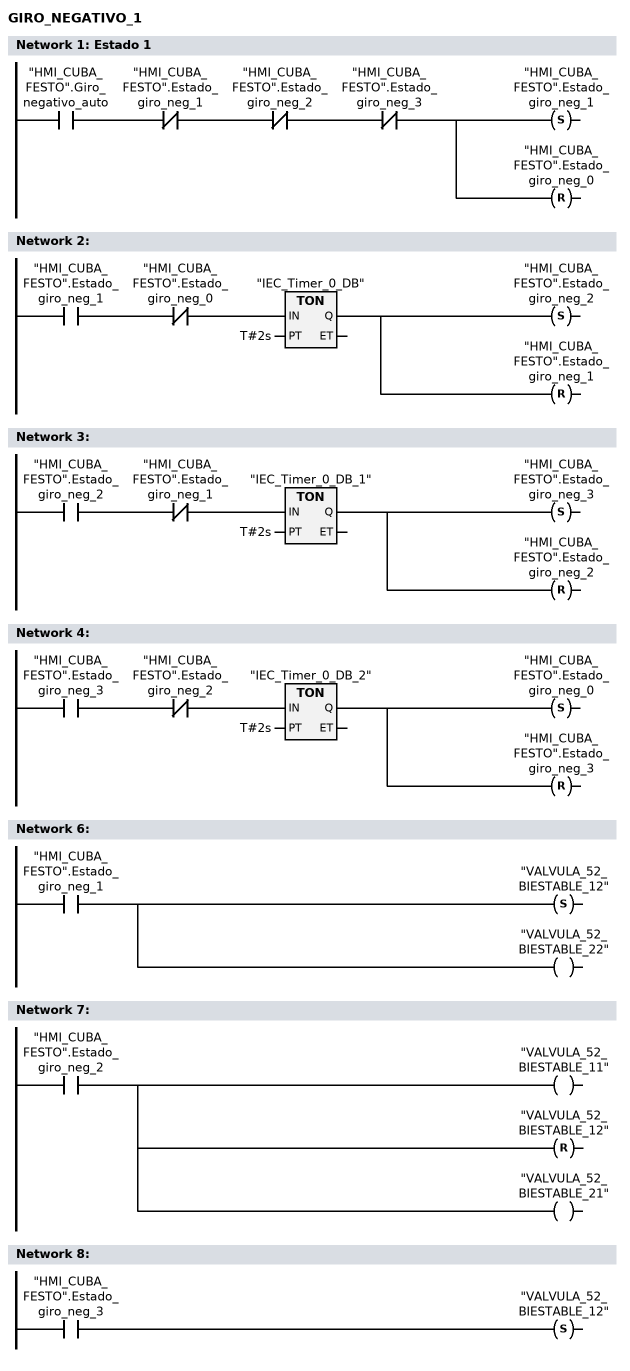
   RUNG wire#powerrail
      Contact( "HMI_CUBA_FESTO".Giro_negativo_auto )
      I_Contact( "HMI_CUBA_FESTO".Estado_giro_neg_1 )
      I_Contact( "HMI_CUBA_FESTO".Estado_giro_neg_2 )
      I_Contact( "HMI_CUBA_FESTO".Estado_giro_neg_3 )
      wire#w1
      S_Coil( "HMI_CUBA_FESTO".Estado_giro_neg_1 )
   END_RUNG
   RUNG wire#w1
      R_Coil( "HMI_CUBA_FESTO".Estado_giro_neg_0 )
   END_RUNG
   // the same network as SCL:
   #_w1 := "HMI_CUBA_FESTO".Giro_negativo_auto AND NOT "HMI_CUBA_FESTO".Estado_giro_neg_1 AND NOT "HMI_CUBA_FESTO".Estado_giro_neg_2 AND NOT "HMI_CUBA_FESTO".Estado_giro_neg_3;
   IF #_w1 THEN
       "HMI_CUBA_FESTO".Estado_giro_neg_1 := TRUE;
       "HMI_CUBA_FESTO".Estado_giro_neg_0 := FALSE;
   END_IF;
END_REGION

REGION Network 2
   "IEC_Timer_0_DB".TON(IN := "HMI_CUBA_FESTO".Estado_giro_neg_1 AND NOT "HMI_CUBA_FESTO".Estado_giro_neg_0,
                        PT := T#2s);
   IF "IEC_Timer_0_DB".Q THEN
       "HMI_CUBA_FESTO".Estado_giro_neg_2 := TRUE;
       "HMI_CUBA_FESTO".Estado_giro_neg_1 := FALSE;
   END_IF;
END_REGION

REGION Network 3
   "IEC_Timer_0_DB_1".TON(IN := "HMI_CUBA_FESTO".Estado_giro_neg_2 AND NOT "HMI_CUBA_FESTO".Estado_giro_neg_1,
                          PT := T#2s);
   IF "IEC_Timer_0_DB_1".Q THEN
       "HMI_CUBA_FESTO".Estado_giro_neg_3 := TRUE;
       "HMI_CUBA_FESTO".Estado_giro_neg_2 := FALSE;
   END_IF;
END_REGION

REGION Network 4
   "IEC_Timer_0_DB_2".TON(IN := "HMI_CUBA_FESTO".Estado_giro_neg_3 AND NOT "HMI_CUBA_FESTO".Estado_giro_neg_2,
                          PT := T#2s);
   IF "IEC_Timer_0_DB_2".Q THEN
       "HMI_CUBA_FESTO".Estado_giro_neg_0 := TRUE;
       "HMI_CUBA_FESTO".Estado_giro_neg_3 := FALSE;
   END_IF;
END_REGION

REGION Network 6
   RUNG wire#powerrail
      Contact( "HMI_CUBA_FESTO".Estado_giro_neg_1 )
      wire#w1
      S_Coil( "VALVULA_52_BIESTABLE_12" )
   END_RUNG
   RUNG wire#w1
      Coil( "VALVULA_52_BIESTABLE_22" )
   END_RUNG
   // the same network as SCL:
   IF "HMI_CUBA_FESTO".Estado_giro_neg_1 THEN "VALVULA_52_BIESTABLE_12" := TRUE; END_IF;
   "VALVULA_52_BIESTABLE_22" := "HMI_CUBA_FESTO".Estado_giro_neg_1;
END_REGION

REGION Network 7
   RUNG wire#powerrail
      Contact( "HMI_CUBA_FESTO".Estado_giro_neg_2 )
      wire#w1
      Coil( "VALVULA_52_BIESTABLE_11" )
   END_RUNG
   RUNG wire#w1
      R_Coil( "VALVULA_52_BIESTABLE_12" )
   END_RUNG
   RUNG wire#w1
      Coil( "VALVULA_52_BIESTABLE_21" )
   END_RUNG
   // the same network as SCL:
   "VALVULA_52_BIESTABLE_11" := "HMI_CUBA_FESTO".Estado_giro_neg_2;
   IF "HMI_CUBA_FESTO".Estado_giro_neg_2 THEN "VALVULA_52_BIESTABLE_12" := FALSE; END_IF;
   "VALVULA_52_BIESTABLE_21" := "HMI_CUBA_FESTO".Estado_giro_neg_2;
END_REGION

REGION Network 8
   RUNG wire#powerrail
      Contact( "HMI_CUBA_FESTO".Estado_giro_neg_3 )
      S_Coil( "VALVULA_52_BIESTABLE_12" )
   END_RUNG
   // the same network as SCL:
   IF "HMI_CUBA_FESTO".Estado_giro_neg_3 THEN "VALVULA_52_BIESTABLE_12" := TRUE; END_IF;
END_REGION
END_FUNCTION_BLOCK

// folder: Achim

FUNCTION_BLOCK "Achim_testPepaFrk"   // FB8, LAD
TITLE = test tools
{ S7_Optimized_Access := 'TRUE' }
VERSION : 0.1
   VAR_INPUT
      inToolIdProxy1 : Bool;
      inToolIdProxy2 : Bool;
      inToolIdProxy3 : Bool;
      inToolIdProxy4 : Bool;
      inAirActivate : Bool;
      inAirPepaCylInActivate : Bool;
      inAirPepaCylOutActivate : Bool;
      inWaterInspPumpActivate : Bool;
      inWaterActivate : Bool;
      inStopRobot : Bool;
      inContRobot : Bool;
      inResetAlarms : Bool;
      inInspRunning : Bool;
      inSTOPMESS : Bool;
      inPRO_ACT : Bool;
      inWaterInspPumpRunning : Bool;
      inWaterInspAlarmFilter : Bool;
      inWaterInspAlarmFc : Bool;
      inWaterInspAlarmElecProt : Bool;
      inWaterInspAlarmUv : Bool;
      inWaterInspAlarmLowLevel : Bool;
      inPepaCylInProxy : Bool;
      inPepaCylOutProxy : Bool;
      inAirOprProxy : Bool;
      inAirMpsCoupledE1 : Bool;
      inAirMpsLockedE2 : Bool;
      inAirMpsUnlockedE3 : Bool;
      inAirMpsPressD1 : Bool;
      inFrkLs1Nc1 : Bool;
      inFrkLs1Nc2 : Bool;
      inFrkLs2Nc1 : Bool;
      inFrkLs2Nc2 : Bool;
      airMpsTimeout : Time := T#500ms;
      airPepaCylTimeout : Time := T#100ms;
      frkLsTimeout : Time := T#100ms;
   END_VAR
   VAR_OUTPUT
      outWaterInspEvL1 : Bool;
      outWaterInspEvL2 : Bool;
      outWaterInspPanelS1 : Bool;
      outWaterInspPanelS2 : Bool;
      outWaterInspPanelS3 : Bool;
      outWaterInspPump : Bool;
      outAirEvOpr : Bool;
      outAirEvMps : Bool;
      outAirPepaCylIn : Bool;
      outAirPepaCylOut : Bool;
      outAntiSpash1 : Bool;
      outAntiSpash2 : Bool;
      outAirMpsAlarm : Bool;
      outAirOprAlarm : Bool;
      outPepaCylAlarm : Bool;
      outFrkLsAlarm : Bool;
      outWaterInspAlarm : Bool;
      outWaterInspAdv : Bool;
      outStopRobot : Bool;
      outMOVE_ENABLE : Bool;
      outCONF_MESS : Bool;
      outEXT_START : Bool;
   END_VAR
   VAR
      tonMpsOn : TON_TIME;
      tonPepaCylOut : TON_TIME;
      tonFrkLs : TON_TIME;
      staticStoppingAlarm : Bool;
      staticAirMpsAlarm : Bool;
      staticAirOprAlarm : Bool;
      staticPepaCylAlarm : Bool;
      staticFrkLsAlarm : Bool;
      staticWaterInspAlarm : Bool;
      staticWaterInspAdv : Bool;
      staticStopRobot : Bool;
      staticContRobot : Bool;
      staticRobotWasStopped : Bool;
      staticairMpsOk : Bool;
      staticTool : Int;
      rtStopRobot : R_TRIG;
      rtContRobot : R_TRIG;
   END_VAR
BEGIN

REGION Network 1 (SCL)
   // tool identification
   IF #inToolIdProxy1 AND NOT #inToolIdProxy2 AND NOT #inToolIdProxy3 AND NOT #inToolIdProxy4 THEN
       #staticTool := 1; // PEPA
   ELSIF NOT #inToolIdProxy1 AND #inToolIdProxy2 AND NOT #inToolIdProxy3 AND NOT #inToolIdProxy4 THEN
       #staticTool := 2; // pole
   ELSIF #inToolIdProxy1 AND #inToolIdProxy2 AND NOT #inToolIdProxy3 AND NOT #inToolIdProxy4 THEN
       #staticTool := 3; // fork
   ELSIF NOT #inToolIdProxy1 AND NOT #inToolIdProxy2 AND #inToolIdProxy3 AND NOT #inToolIdProxy4 THEN
       #staticTool := 4; // teaching
   ELSIF #inToolIdProxy1 AND NOT #inToolIdProxy2 AND #inToolIdProxy3 AND NOT #inToolIdProxy4 THEN
       #staticTool := 5; // marker    
   ELSIF NOT #inToolIdProxy1 AND NOT #inToolIdProxy2 AND NOT #inToolIdProxy3 AND NOT #inToolIdProxy4 THEN
       #staticTool := 0; // no tool  
   ELSE
       #staticTool := -1; // unknown
   END_IF;

   // air MPS & OPR activation
   #outAirEvOpr := #inAirActivate AND (#staticTool=1 OR #staticTool=2 OR #staticTool=5);
   #outAirEvMps := #inAirActivate;

   // check MPS & OPR signals
   #staticairMpsOk := #inAirMpsCoupledE1 AND #inAirMpsLockedE2 AND NOT #inAirMpsUnlockedE3 AND #inAirMpsPressD1;
   #tonMpsOn(IN := #inAirActivate AND #staticTool>0,
                 PT := #airMpsTimeout);
   IF #tonMpsOn.Q THEN
           IF NOT #staticairMpsOk THEN
               #staticAirMpsAlarm := true;
           END_IF;
           IF NOT #inAirOprProxy AND (#staticTool=1 OR #staticTool=2 OR #staticTool=5) THEN
               #staticAirOprAlarm := true;
           END_IF;
   END_IF;

   // alarms
   IF #inResetAlarms THEN
       #staticAirMpsAlarm := false;
       #staticAirOprAlarm := false;
       #staticPepaCylAlarm := false;
       #staticFrkLsAlarm := false;
       #staticWaterInspAlarm := false;
       #staticWaterInspAdv := false;
   END_IF;
   IF #inResetAlarms AND #inSTOPMESS THEN
       #outCONF_MESS := true;
   ELSE
       #outCONF_MESS := false;
   END_IF;

   #rtContRobot(CLK := #inContRobot);
   IF #staticRobotWasStopped AND #rtContRobot.Q AND NOT #staticStoppingAlarm THEN
       #staticContRobot := true;
       #staticRobotWasStopped := false;
   END_IF;

   // water pump
   IF #inWaterInspAlarmFilter OR #inWaterInspAlarmUv THEN
       #staticWaterInspAdv := true;
   END_IF;
   IF (#inWaterInspAlarmFc OR #inWaterInspAlarmElecProt OR #inWaterInspAlarmLowLevel) AND #inWaterActivate THEN
       #staticWaterInspAlarm := true;
   END_IF;
   #outWaterInspPump := #inWaterInspPumpActivate AND NOT #staticWaterInspAlarm;

   // water valves
   #outWaterInspPanelS1 := #inWaterActivate AND #inWaterInspPumpRunning AND #staticTool=3;
   #outWaterInspPanelS2 := #inWaterActivate AND #inWaterInspPumpRunning AND #staticTool=3;
   #outWaterInspPanelS3 := #inWaterActivate AND #inWaterInspPumpRunning AND #staticTool=1;
   #outWaterInspEvL1 := #inWaterActivate AND #inWaterInspPumpRunning AND #staticTool = 3;
   #outWaterInspEvL2 := #inWaterActivate AND #inWaterInspPumpRunning AND (#staticTool=1 OR #staticTool=3);

   // retract & extend PEPA / marker cylinder
   #outAirPepaCylIn := #inAirPepaCylInActivate AND (#staticTool=1 OR #staticTool=5);
   #outAirPepaCylOut := #inAirPepaCylOutActivate AND (#staticTool=1 OR #staticTool=5);

   // anti splash air FRK
   #outAntiSpash1 := #inInspRunning AND #staticTool=3;
   #outAntiSpash2 := #inInspRunning AND #staticTool=3;

   // check micro cyl in / cyl out triggers while PEPA cyl out during inspection
   #tonPepaCylOut(IN := #inInspRunning AND (#inPepaCylInProxy OR #inPepaCylOutProxy) AND (#staticTool=1 OR #staticTool=5),
                       PT := #airPepaCylTimeout);
   IF #tonPepaCylOut.Q THEN
       #staticPepaCylAlarm := true;
   END_IF;

   // check limit switches FRK
   #tonFrkLs(IN := (NOT #inFrkLs1Nc1 OR NOT #inFrkLs1Nc2 OR NOT #inFrkLs2Nc1 OR NOT #inFrkLs2Nc1 OR NOT #inFrkLs2Nc2) AND #staticTool=3,
             PT := #frkLsTimeout);
   IF #tonFrkLs.Q THEN
       #staticFrkLsAlarm := true;
   END_IF;

   // stop robot
   #staticStoppingAlarm := #staticAirMpsAlarm OR #staticAirOprAlarm OR #staticWaterInspAlarm OR #staticPepaCylAlarm OR #staticFrkLsAlarm;
   #rtStopRobot(CLK := #inStopRobot OR #staticStoppingAlarm);
   IF #rtStopRobot.Q THEN
       #staticStopRobot := true;
   END_IF;

   // feedback stop robot cmd from robot
   IF #staticStopRobot AND #inSTOPMESS AND NOT #inPRO_ACT THEN
       #staticStopRobot := false;
       #staticRobotWasStopped := true;
   END_IF;

   // feedback cont robot cmd from robot
   IF #staticContRobot AND #inPRO_ACT THEN
       #staticContRobot := false;
   END_IF;

   // outputs
   #outStopRobot := #staticStopRobot;
   #outMOVE_ENABLE := NOT #staticStopRobot;
   #outEXT_START := #staticContRobot;
   #outAirMpsAlarm := #staticAirMpsAlarm;
   #outAirOprAlarm := #staticAirOprAlarm;
   #outPepaCylAlarm := #staticPepaCylAlarm;
   #outFrkLsAlarm := #staticFrkLsAlarm;
   #outWaterInspAlarm := #staticWaterInspAlarm;
   #outWaterInspAdv := #staticWaterInspAdv;
END_REGION
END_FUNCTION_BLOCK

FUNCTION "Achim" : Void   // FC1, LAD
{ S7_Optimized_Access := 'TRUE' }
VERSION : 0.1
BEGIN

REGION Network 1: test end effector
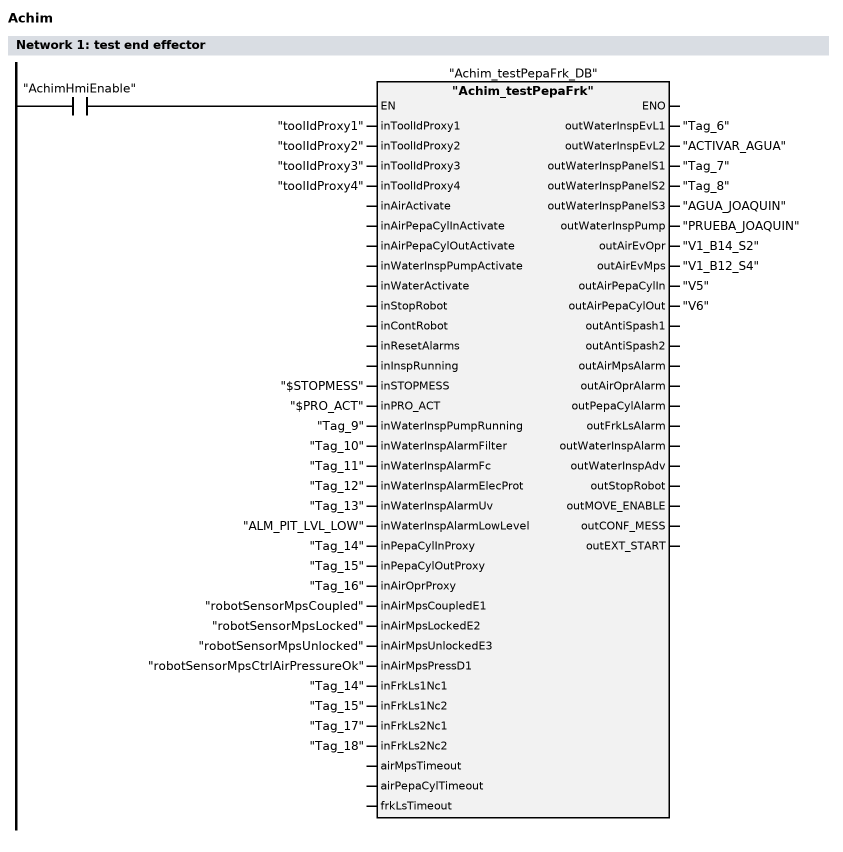
   RUNG wire#powerrail
      Contact( "AchimHmiEnable" )
      "Achim_testPepaFrk_DB"(inToolIdProxy1 := "toolIdProxy1", inToolIdProxy2 := "toolIdProxy2", inToolIdProxy3 := "toolIdProxy3", inToolIdProxy4 := "toolIdProxy4", inAirActivate :=, inAirPepaCylInActivate :=, inAirPepaCylOutActivate :=, inWaterInspPumpActivate :=, inWaterActivate :=, inStopRobot :=, inContRobot :=, inResetAlarms :=, inInspRunning :=, inSTOPMESS := "$STOPMESS", inPRO_ACT := "$PRO_ACT", inWaterInspPumpRunning := "Tag_9", inWaterInspAlarmFilter := "Tag_10", inWaterInspAlarmFc := "Tag_11", inWaterInspAlarmElecProt := "Tag_12", inWaterInspAlarmUv := "Tag_13", inWaterInspAlarmLowLevel := "ALM_PIT_LVL_LOW", inPepaCylInProxy := "Tag_14", inPepaCylOutProxy := "Tag_15", inAirOprProxy := "Tag_16", inAirMpsCoupledE1 := "robotSensorMpsCoupled", inAirMpsLockedE2 := "robotSensorMpsLocked", inAirMpsUnlockedE3 := "robotSensorMpsUnlocked", inAirMpsPressD1 := "robotSensorMpsCtrlAirPressureOk", inFrkLs1Nc1 := "Tag_14", inFrkLs1Nc2 := "Tag_15", inFrkLs2Nc1 := "Tag_17", inFrkLs2Nc2 := "Tag_18", airMpsTimeout :=, airPepaCylTimeout :=, frkLsTimeout :=, outWaterInspEvL1 => "Tag_6", outWaterInspEvL2 => "ACTIVAR_AGUA", outWaterInspPanelS1 => "Tag_7", outWaterInspPanelS2 => "Tag_8", outWaterInspPanelS3 => "AGUA_JOAQUIN", outWaterInspPump => "PRUEBA_JOAQUIN", outAirEvOpr => "V1_B14_S2", outAirEvMps => "V1_B12_S4", outAirPepaCylIn => "V5", outAirPepaCylOut => "V6", outAntiSpash1 =>, outAntiSpash2 =>, outAirMpsAlarm =>, outAirOprAlarm =>, outPepaCylAlarm =>, outFrkLsAlarm =>, outWaterInspAlarm =>, outWaterInspAdv =>, outStopRobot =>, outMOVE_ENABLE =>, outCONF_MESS =>, outEXT_START =>)
   END_RUNG
   // the same network as SCL:
   IF "AchimHmiEnable" THEN
       "Achim_testPepaFrk_DB"(inToolIdProxy1 := "toolIdProxy1",   // "Achim_testPepaFrk"
                              inToolIdProxy2 := "toolIdProxy2",
                              inToolIdProxy3 := "toolIdProxy3",
                              inToolIdProxy4 := "toolIdProxy4",
                              inSTOPMESS := "$STOPMESS",
                              inPRO_ACT := "$PRO_ACT",
                              inWaterInspPumpRunning := "Tag_9",
                              inWaterInspAlarmFilter := "Tag_10",
                              inWaterInspAlarmFc := "Tag_11",
                              inWaterInspAlarmElecProt := "Tag_12",
                              inWaterInspAlarmUv := "Tag_13",
                              inWaterInspAlarmLowLevel := "ALM_PIT_LVL_LOW",
                              inPepaCylInProxy := "Tag_14",
                              inPepaCylOutProxy := "Tag_15",
                              inAirOprProxy := "Tag_16",
                              inAirMpsCoupledE1 := "robotSensorMpsCoupled",
                              inAirMpsLockedE2 := "robotSensorMpsLocked",
                              inAirMpsUnlockedE3 := "robotSensorMpsUnlocked",
                              inAirMpsPressD1 := "robotSensorMpsCtrlAirPressureOk",
                              inFrkLs1Nc1 := "Tag_14",
                              inFrkLs1Nc2 := "Tag_15",
                              inFrkLs2Nc1 := "Tag_17",
                              inFrkLs2Nc2 := "Tag_18",
                              outWaterInspEvL1 => "Tag_6",
                              outWaterInspEvL2 => "ACTIVAR_AGUA",
                              outWaterInspPanelS1 => "Tag_7",
                              outWaterInspPanelS2 => "Tag_8",
                              outWaterInspPanelS3 => "AGUA_JOAQUIN",
                              outWaterInspPump => "PRUEBA_JOAQUIN",
                              outAirEvOpr => "V1_B14_S2",
                              outAirEvMps => "V1_B12_S4",
                              outAirPepaCylIn => "V5",
                              outAirPepaCylOut => "V6");
   END_IF;
END_REGION
END_FUNCTION

(* ===== HMI "HMI_RT_1" =====
system functions are stored by id; their names below are inferred from use
connection "HMI_Connection_1": ETHERNET, SMART_S7_1200_OMS

HMI tags "Default tag table"
   "Tag_ScreenNumber" : UInt, internal

HMI tags "CUBA_FESTO"
   "HMI_CUBA_FESTO_HMI_Sensor_plato_giro_1" : Bool = PLC HMI_CUBA_FESTO.HMI_Sensor_plato_giro_1, 100 ms
   "HMI_CUBA_FESTO_HMI_Sensor_Plato_giro_2" : Bool = PLC HMI_CUBA_FESTO.HMI_Sensor_Plato_giro_2, 100 ms
   "HMI_CUBA_FESTO_HMI_Sensor_plato_giro_3" : Bool = PLC HMI_CUBA_FESTO.HMI_Sensor_plato_giro_3, 100 ms
   "HMI_CUBA_FESTO_HMI_Sensor_ADN_bastidor_bloqueado_1" : Bool = PLC HMI_CUBA_FESTO.HMI_Sensor_ADN_bastidor_bloqueado_1, 100 ms
   "HMI_CUBA_FESTO_HMI_Sensor_ADN_bastidor_desbloqueado_1" : Bool = PLC HMI_CUBA_FESTO.HMI_Sensor_ADN_bastidor_desbloqueado_1, 100 ms
   "HMI_CUBA_FESTO_HMI_Sensor_ADN_bastidor_bloqueado_2" : Bool = PLC HMI_CUBA_FESTO.HMI_Sensor_ADN_bastidor_bloqueado_2, 100 ms
   "HMI_CUBA_FESTO_HMI_Sensor_ADN_bastidor_desbloqueado_2" : Bool = PLC HMI_CUBA_FESTO.HMI_Sensor_ADN_bastidor_desbloqueado_2, 100 ms
   "HMI_CUBA_FESTO_HMI_SENSOR_CRDSNU_BASTIDOR_BLOQUEADO_1" : Bool = PLC HMI_CUBA_FESTO.HMI_SENSOR_CRDSNU_BASTIDOR_BLOQUEADO_1, 100 ms
   "HMI_CUBA_FESTO_HMI_SENSOR_CRDSNU_BASTIDOR_DESBLOQUEADO_1" : Bool = PLC HMI_CUBA_FESTO.HMI_SENSOR_CRDSNU_BASTIDOR_DESBLOQUEADO_1, 100 ms
   "HMI_CUBA_FESTO_HMI_SENSOR_CRDSNU_BASTIDOR_BLOQUEADO_2" : Bool = PLC HMI_CUBA_FESTO.HMI_SENSOR_CRDSNU_BASTIDOR_BLOQUEADO_2, 100 ms
   "HMI_CUBA_FESTO_HMI_SENSOR_CRDSNU_BASTIDOR_DESBLOQUEADO_2" : Bool = PLC HMI_CUBA_FESTO.HMI_SENSOR_CRDSNU_BASTIDOR_DESBLOQUEADO_2, 100 ms
   "HMI_CUBA_FESTO_HMI_SENSOR_DSBG_BASTIDOR_ARRIBA_1" : Bool = PLC HMI_CUBA_FESTO.HMI_SENSOR_DSBG_BASTIDOR_ARRIBA_1, 100 ms
   "HMI_CUBA_FESTO_HMI_SENSOR_DSBG_BASTIDOR_ABAJO_1" : Bool = PLC HMI_CUBA_FESTO.HMI_SENSOR_DSBG_BASTIDOR_ABAJO_1, 100 ms
   "HMI_CUBA_FESTO_HMI_SENSOR_DSBG_BASTIDOR_ARRIBA_2" : Bool = PLC HMI_CUBA_FESTO.HMI_SENSOR_DSBG_BASTIDOR_ARRIBA_2, 100 ms
   "HMI_CUBA_FESTO_HMI_SENSOR_DSBG_BASTIDOR_ABAJO_2" : Bool = PLC HMI_CUBA_FESTO.HMI_SENSOR_DSBG_BASTIDOR_ABAJO_2, 100 ms
   "HMI_CUBA_FESTO_HMI_PULSADOR_SUBIR_1" : Bool = PLC HMI_CUBA_FESTO.HMI_PULSADOR_SUBIR_1, 100 ms
   "HMI_CUBA_FESTO_HMI_PULSADOR_BAJAR_1" : Bool = PLC HMI_CUBA_FESTO.HMI_PULSADOR_BAJAR_1, 100 ms
   "HMI_CUBA_FESTO_HMI_PULSADOR_SUBIR_2" : Bool = PLC HMI_CUBA_FESTO.HMI_PULSADOR_SUBIR_2, 100 ms
   "HMI_CUBA_FESTO_HMI_PULSADOR_BAJAR_2" : Bool = PLC HMI_CUBA_FESTO.HMI_PULSADOR_BAJAR_2, 100 ms
   "HMI_CUBA_FESTO_HMI_VALVULA_52_BIESTABLE_11" : Bool = PLC HMI_CUBA_FESTO.HMI_VALVULA_52_BIESTABLE_11, 100 ms
   "HMI_CUBA_FESTO_HMI_VALVULA_52_BIESTABLE_12" : Bool = PLC HMI_CUBA_FESTO.HMI_VALVULA_52_BIESTABLE_12, 100 ms
   "HMI_CUBA_FESTO_HMI_VALVULA_52_BIESTABLE_21" : Bool = PLC HMI_CUBA_FESTO.HMI_VALVULA_52_BIESTABLE_21 AT %DB1.DBX0.0, 100 ms
   "HMI_CUBA_FESTO_HMI_VALVULA_52_BIESTABLE_22" : Bool = PLC HMI_CUBA_FESTO.HMI_VALVULA_52_BIESTABLE_22 AT %DB1.DBX0.0, 100 ms
   "HMI_CUBA_FESTO_HMI_VÁLVULA_52_MONOESTABLE_1" : Bool = PLC HMI_CUBA_FESTO.HMI_VÁLVULA_52_MONOESTABLE_1 AT %DB1.DBX0.0, 100 ms
   "HMI_CUBA_FESTO_HMI_VÁLVULA_52_MONOESTABLE_2" : Bool = PLC HMI_CUBA_FESTO.HMI_VÁLVULA_52_MONOESTABLE_2 AT %DB1.DBX0.0, 100 ms
   "HMI_CUBA_FESTO_HMI_VÁLVULA_52_MONOESTABLE_3" : Bool = PLC HMI_CUBA_FESTO.HMI_VÁLVULA_52_MONOESTABLE_3 AT %DB1.DBX0.0, 100 ms
   "HMI_CUBA_FESTO_HMI_VÁLVULA_52_MONOESTABLE_4" : Bool = PLC HMI_CUBA_FESTO.HMI_VÁLVULA_52_MONOESTABLE_4 AT %DB1.DBX0.0, 100 ms
   "HMI_CUBA_FESTO_HMI_VÁLVULA_52_MONOESTABLE_5" : Bool = PLC HMI_CUBA_FESTO.HMI_VÁLVULA_52_MONOESTABLE_5 AT %DB1.DBX0.0, 100 ms
   "HMI_CUBA_FESTO_HMI_VÁLVULA_52_MONOESTABLE_6" : Bool = PLC HMI_CUBA_FESTO.HMI_VÁLVULA_52_MONOESTABLE_6 AT %DB1.DBX0.0, 100 ms
   "HMI_CUBA_FESTO_HMI_VÁLVULA_52_MONOESTABLE_7" : Bool = PLC HMI_CUBA_FESTO.HMI_VÁLVULA_52_MONOESTABLE_7 AT %DB1.DBX0.0, 100 ms
   "HMI_CUBA_FESTO_HMI_VÁLVULA_52_MONOESTABLE_8" : Bool = PLC HMI_CUBA_FESTO.HMI_VÁLVULA_52_MONOESTABLE_8 AT %DB1.DBX0.0, 100 ms
   "HMI_CUBA_FESTO_HMI_VÁLVULA_52_MONOESTABLE_9" : Bool = PLC HMI_CUBA_FESTO.HMI_VÁLVULA_52_MONOESTABLE_9 AT %DB1.DBX0.0, 100 ms
   "HMI_CUBA_FESTO_HMI_VÁLVULA_52_MONOESTABLE_10" : Bool = PLC HMI_CUBA_FESTO.HMI_VÁLVULA_52_MONOESTABLE_10 AT %DB1.DBX0.0, 100 ms
   "HMI_CUBA_FESTO_HMI_VÁLVULA_52_MONOESTABLE_11" : Bool = PLC HMI_CUBA_FESTO.HMI_VÁLVULA_52_MONOESTABLE_11 AT %DB1.DBX0.0, 100 ms
   "HMI_CUBA_FESTO_HMI_VÁLVULA_52_MONOESTABLE_12" : Bool = PLC HMI_CUBA_FESTO.HMI_VÁLVULA_52_MONOESTABLE_12 AT %DB1.DBX0.0, 100 ms
   "HMI_CUBA_FESTO_HMI_VÁLVULA_52_MONOESTABLE_13" : Bool = PLC HMI_CUBA_FESTO.HMI_VÁLVULA_52_MONOESTABLE_13 AT %DB1.DBX0.0, 100 ms
   "HMI_CUBA_FESTO_HMI_VÁLVULA_52_MONOESTABLE_14" : Bool = PLC HMI_CUBA_FESTO.HMI_VÁLVULA_52_MONOESTABLE_14 AT %DB1.DBX0.0, 100 ms
   "HMI_CUBA_FESTO_HMI_VÁLVULA_52_MONOESTABLE_15" : Bool = PLC HMI_CUBA_FESTO.HMI_VÁLVULA_52_MONOESTABLE_15 AT %DB1.DBX0.0, 100 ms
   "HMI_CUBA_FESTO_HMI_VÁLVULA_52_MONOESTABLE_16" : Bool = PLC HMI_CUBA_FESTO.HMI_VÁLVULA_52_MONOESTABLE_16 AT %DB1.DBX0.0, 100 ms
   "HMI_CUBA_FESTO_HMI_VÁLVULA_52_MONOESTABLE_17" : Bool = PLC HMI_CUBA_FESTO.HMI_VÁLVULA_52_MONOESTABLE_17 AT %DB1.DBX0.0, 100 ms
   "HMI_CUBA_FESTO_HMI_VÁLVULA_52_MONOESTABLE_18" : Bool = PLC HMI_CUBA_FESTO.HMI_VÁLVULA_52_MONOESTABLE_18 AT %DB1.DBX0.0, 100 ms
   "HMI_CUBA_FESTO_HMI_VÁLVULA_52_MONOESTABLE_19" : Bool = PLC HMI_CUBA_FESTO.HMI_VÁLVULA_52_MONOESTABLE_19 AT %DB1.DBX0.0, 100 ms
   "HMI_CUBA_FESTO_HMI_VÁLVULA_52_MONOESTABLE_20" : Bool = PLC HMI_CUBA_FESTO.HMI_VÁLVULA_52_MONOESTABLE_20 AT %DB1.DBX0.0, 100 ms
   "HMI_CUBA_FESTO_HMI_VÁLVULA_52_MONOESTABLE_21" : Bool = PLC HMI_CUBA_FESTO.HMI_VÁLVULA_52_MONOESTABLE_21 AT %DB1.DBX0.0, 100 ms
   "HMI_CUBA_FESTO_HMI_VÁLVULA_52_MONOESTABLE_22" : Bool = PLC HMI_CUBA_FESTO.HMI_VÁLVULA_52_MONOESTABLE_22 AT %DB1.DBX0.0, 100 ms
   "HMI_CUBA_FESTO_HMI_VÁLVULA_52_MONOESTABLE_23" : Bool = PLC HMI_CUBA_FESTO.HMI_VÁLVULA_52_MONOESTABLE_23 AT %DB1.DBX0.0, 100 ms
   "HMI_CUBA_FESTO_HMI_VÁLVULA_52_MONOESTABLE_24" : Bool = PLC HMI_CUBA_FESTO.HMI_VÁLVULA_52_MONOESTABLE_24 AT %DB1.DBX0.0, 100 ms
   "HMI_CUBA_FESTO_HMI_VÁLVULA_52_MONOESTABLE_25" : Bool = PLC HMI_CUBA_FESTO.HMI_VÁLVULA_52_MONOESTABLE_25 AT %DB1.DBX0.0, 100 ms
   "HMI_CUBA_FESTO_HMI_VÁLVULA_52_MONOESTABLE_26" : Bool = PLC HMI_CUBA_FESTO.HMI_VÁLVULA_52_MONOESTABLE_26 AT %DB1.DBX0.0, 100 ms
   "HMI_CUBA_FESTO_HMI_VÁLVULA_52_MONOESTABLE_27" : Bool = PLC HMI_CUBA_FESTO.HMI_VÁLVULA_52_MONOESTABLE_27 AT %DB1.DBX0.0, 100 ms
   "HMI_CUBA_FESTO_HMI_VÁLVULA_52_MONOESTABLE_28" : Bool = PLC HMI_CUBA_FESTO.HMI_VÁLVULA_52_MONOESTABLE_28 AT %DB1.DBX0.0, 100 ms
   "HMI_CUBA_FESTO_HMI_PULSADOR_BAJAR_3" : Bool = PLC HMI_CUBA_FESTO.HMI_PULSADOR_BAJAR_3 AT %DB1.DBX0.0, 100 ms
   "HMI_CUBA_FESTO_HMI_PULSADOR_BAJAR_4" : Bool = PLC HMI_CUBA_FESTO.HMI_PULSADOR_BAJAR_4 AT %DB1.DBX0.0, 100 ms
   "HMI_CUBA_FESTO_HMI_PULSADOR_BAJAR_5" : Bool = PLC HMI_CUBA_FESTO.HMI_PULSADOR_BAJAR_5 AT %DB1.DBX0.0, 100 ms
   "HMI_CUBA_FESTO_HMI_PULSADOR_BAJAR_6" : Bool = PLC HMI_CUBA_FESTO.HMI_PULSADOR_BAJAR_6 AT %DB1.DBX0.0, 100 ms
   "HMI_CUBA_FESTO_HMI_PULSADOR_BAJAR_7" : Bool = PLC HMI_CUBA_FESTO.HMI_PULSADOR_BAJAR_7 AT %DB1.DBX0.0, 100 ms
   "HMI_CUBA_FESTO_HMI_PULSADOR_BAJAR_8" : Bool = PLC HMI_CUBA_FESTO.HMI_PULSADOR_BAJAR_8 AT %DB1.DBX0.0, 100 ms
   "HMI_CUBA_FESTO_HMI_PULSADOR_BAJAR_9" : Bool = PLC HMI_CUBA_FESTO.HMI_PULSADOR_BAJAR_9 AT %DB1.DBX0.0, 100 ms
   "HMI_CUBA_FESTO_HMI_PULSADOR_BAJAR_10" : Bool = PLC HMI_CUBA_FESTO.HMI_PULSADOR_BAJAR_10 AT %DB1.DBX0.0, 100 ms
   "HMI_CUBA_FESTO_HMI_PULSADOR_BAJAR_11" : Bool = PLC HMI_CUBA_FESTO.HMI_PULSADOR_BAJAR_11 AT %DB1.DBX0.0, 100 ms
   "HMI_CUBA_FESTO_HMI_PULSADOR_BAJAR_12" : Bool = PLC HMI_CUBA_FESTO.HMI_PULSADOR_BAJAR_12 AT %DB1.DBX0.0, 100 ms
   "HMI_CUBA_FESTO_HMI_PULSADOR_BAJAR_13" : Bool = PLC HMI_CUBA_FESTO.HMI_PULSADOR_BAJAR_13 AT %DB1.DBX0.0, 100 ms
   "HMI_CUBA_FESTO_HMI_PULSADOR_BAJAR_14" : Bool = PLC HMI_CUBA_FESTO.HMI_PULSADOR_BAJAR_14 AT %DB1.DBX0.0, 100 ms
   "HMI_CUBA_FESTO_HMI_HABILITAR_AUTOMATICO" : Bool = PLC HMI_CUBA_FESTO.GIRO_AUTOMATICO_HABILITADO AT %DB1.DBX0.0, 1 s
   "HMI_CUBA_FESTO_HMI_GIRO_POSITIVO_AUTO" : Bool = PLC HMI_CUBA_FESTO.Giro_positivo_auto AT %DB1.DBX0.0, 1 s
   "HMI_CUBA_FESTO_HMI_GIRO_NEGATIVO_AUTO" : Bool = PLC HMI_CUBA_FESTO.Giro_negativo_auto AT %DB1.DBX0.0, 1 s

HMI tags "Achim_test"
   "hmiAchimAir" : Bool = PLC Achim_testPepaFrk_DB.inAirActivate AT %DB1.DBX0.0, 1 s
   "hmiAchimPepaCylIn" : Bool = PLC Achim_testPepaFrk_DB.inAirPepaCylInActivate AT %DB1.DBX0.0, 1 s
   "hmiAchimPepaCylOut" : Bool = PLC Achim_testPepaFrk_DB.inAirPepaCylOutActivate AT %DB1.DBX0.0, 1 s
   "hmiAchimWaterInspPump" : Bool = PLC Achim_testPepaFrk_DB.inWaterInspPumpActivate AT %DB1.DBX0.0, 1 s
   "hmiAchimWaterActivate" : Bool = PLC Achim_testPepaFrk_DB.inWaterActivate AT %DB1.DBX0.0, 1 s
   "hmiAchimStopRobot" : Bool = PLC Achim_testPepaFrk_DB.inStopRobot AT %DB1.DBX0.0, 1 s
   "hmiAchimContRobot" : Bool = PLC Achim_testPepaFrk_DB.inContRobot AT %DB1.DBX0.0, 1 s
   "hmiAchimResetAlarms" : Bool = PLC Achim_testPepaFrk_DB.inResetAlarms AT %DB1.DBX0.0, 1 s
   "hmiAchimInspRunning" : Bool = PLC Achim_testPepaFrk_DB.inInspRunning AT %DB1.DBX0.0, 1 s
   "hmiAchimWaterInspPumpRunning" : Bool = PLC Achim_testPepaFrk_DB.inWaterInspPumpRunning AT %DB1.DBX0.0, 1 s
   "hmiAchimWaterL1" : Bool = PLC Achim_testPepaFrk_DB.outWaterInspEvL1 AT %DB1.DBX0.0, 1 s
   "hmiAchimWaterL2" : Bool = PLC Achim_testPepaFrk_DB.outWaterInspEvL2 AT %DB1.DBX0.0, 1 s
   "hmiAchimWaterS1" : Bool = PLC Achim_testPepaFrk_DB.outWaterInspPanelS1 AT %DB1.DBX0.0, 1 s
   "hmiAchimWaterS2" : Bool = PLC Achim_testPepaFrk_DB.outWaterInspPanelS2 AT %DB1.DBX0.0, 1 s
   "hmiAchimWaterS3" : Bool = PLC Achim_testPepaFrk_DB.outWaterInspPanelS3 AT %DB1.DBX0.0, 1 s
   "hmiAchimMpsEv" : Bool = PLC Achim_testPepaFrk_DB.outAirEvMps AT %DB1.DBX0.0, 1 s
   "hmiAchimOprEv" : Bool = PLC Achim_testPepaFrk_DB.outAirEvOpr AT %DB1.DBX0.0, 1 s
   "hmiAchimAntiSpash" : Bool = PLC Achim_testPepaFrk_DB.outAntiSpash1 AT %DB1.DBX0.0, 1 s
   "hmiAchimMpsAlarm" : Bool = PLC Achim_testPepaFrk_DB.outAirMpsAlarm AT %DB1.DBX0.0, 1 s
   "hmiAchimOprAlarm" : Bool = PLC Achim_testPepaFrk_DB.outAirOprAlarm AT %DB1.DBX0.0, 1 s
   "hmiAchimPepaCylAlarm" : Bool = PLC Achim_testPepaFrk_DB.outPepaCylAlarm AT %DB1.DBX0.0, 1 s
   "hmiAchimFrkLsAlarm" : Bool = PLC Achim_testPepaFrk_DB.outFrkLsAlarm AT %DB1.DBX0.0, 1 s
   "hmiAchimWaterInspAlarm" : Bool = PLC Achim_testPepaFrk_DB.outWaterInspAlarm AT %DB1.DBX0.0, 1 s
   "hmiAchimWaterInspAdv" : Bool = PLC Achim_testPepaFrk_DB.outWaterInspAdv AT %DB1.DBX0.0, 1 s
   "hmiAchimAirMpsCoupledE1" : Bool = PLC Achim_testPepaFrk_DB.inAirMpsCoupledE1 AT %DB1.DBX0.0, 1 s
   "hmiAchimAirMpsLockedE2" : Bool = PLC Achim_testPepaFrk_DB.inAirMpsLockedE2 AT %DB1.DBX0.0, 1 s
   "hmiAchimAirMpsUnlockedE3" : Bool = PLC Achim_testPepaFrk_DB.inAirMpsUnlockedE3 AT %DB1.DBX0.0, 1 s
   "hmiAchimAirMpsPressD1" : Bool = PLC Achim_testPepaFrk_DB.inAirMpsPressD1 AT %DB1.DBX0.0, 1 s
   "hmiAchimPepaCylInProxy" : Bool = PLC Achim_testPepaFrk_DB.inPepaCylInProxy AT %DB1.DBX0.0, 1 s
   "hmiAchimPepaCylOutProxy" : Bool = PLC Achim_testPepaFrk_DB.inPepaCylOutProxy AT %DB1.DBX0.0, 1 s
   "hmiAchimFrkLs1Nc1" : Bool = PLC Achim_testPepaFrk_DB.inFrkLs1Nc1 AT %DB1.DBX0.0, 1 s
   "hmiAchimFrkLs1Nc2" : Bool = PLC Achim_testPepaFrk_DB.inFrkLs1Nc2 AT %DB1.DBX0.0, 1 s
   "hmiAchimFrkLs2Nc1" : Bool = PLC Achim_testPepaFrk_DB.inFrkLs2Nc1 AT %DB1.DBX0.0, 1 s
   "hmiAchimFrkLs2Nc2" : Bool = PLC Achim_testPepaFrk_DB.inFrkLs2Nc2 AT %DB1.DBX0.0, 1 s
   "hmiAchimOprProxy" : Bool = PLC Achim_testPepaFrk_DB.inAirOprProxy AT %DB1.DBX0.0, 1 s
   "hmiAchimEnable" : Bool = PLC AchimHmiEnable AT %M202.0, 1 s
   "hmiAchimTool" : Int = PLC Achim_testPepaFrk_DB.staticTool AT %DB1.DBX0.0, 1 s
   "hmiAchimSTOPMESS" : Bool = PLC Achim_testPepaFrk_DB.inSTOPMESS AT %DB1.DBX0.0, 1 s
   "hmiAchimPRO_ACT" : Bool = PLC Achim_testPepaFrk_DB.inPRO_ACT AT %DB1.DBX0.0, 1 s

text list "tool": -1 'unknown'; 0 'no tool'; 1 'PEPA'; 2 'pole'; 3 'yugo'; 4 'teaching'; 5 'marcador'

Template "Template_1" 1280x800
   Button "Exit" at 1182,752 size 67x47; TextOff 'Exit'; PictureOff "ExitRuntime_KTP1200_Basic_PN_TR"; PictureOn "ExitRuntime_KTP1200_Basic_PN_TR"
      on Release: StopRuntime(0)
   Button "Template_Button" at 1054,752 size 67x47; TextOff 'Text'
   Button "Template_Button_1" at 926,752 size 67x47; TextOff 'Text'
   Button "Template_Button_2" at 798,752 size 67x47; TextOff 'Text'
   Button "Template_Button_3" at 670,752 size 67x47; TextOff 'Text'
   Button "Template_Button_4" at 542,752 size 67x47; TextOff 'Text'
   Button "Template_Button_5" at 414,752 size 67x47; TextOff 'Text'
   Button "Template_Button_6" at 286,752 size 67x47; TextOff 'Text'
   Button "Alarms" at 158,752 size 67x47; TextOff 'Alarms'; PictureOff "AlarmDisplay_KTP1200_Basic_PN_TR"; PictureOn "AlarmDisplay_KTP1200_Basic_PN_TR"
      on Release: function_ef3f5d25("Alarm window_Unacknowledged", -1)
   Button "Start screen" at 30,752 size 67x47; TextOff 'Start screen'; PictureOff "NavigateHome_KTP1200_Basic_PN_TR"; PictureOn "NavigateHome_KTP1200_Basic_PN_TR"
      on Release: ActivateScreen("Root screen", 0)
   SymbolicIOField "Symbolic_IO_Field_Screen" at 87,9 size 1086x30; TextOff '0'; TextOn '1'; TextList "TextList_ScreenNames"
      ProcessValue <- "Tag_ScreenNumber"
      on Change: ActivateScreenByNumber("Tag_ScreenNumber", 0)
   DateTimeField "HmiScreenItemData" at 1175,24 size 105x24
   DateTimeField "HmiScreenItemData_1" at 1175,0 size 105x24
   GraphicView "Logo" at 0,0 size 85x48; Picture "Logo of HMI_1"

screen "Root screen" 1280x800, template "Template_1"
   on GenerateScreen: SetTag("Tag_ScreenNumber", 1)
   TextField "HmiScreenItemData_1" at 128,384 size 1024x27; Text 'Welcome to HMI_1 (KTP1200 Basic+ PN)!'
   Button "HmiScreenItemData" at 36,84 size 159x47; TextOff 'Screen_Prueba'; PictureOff "Navigates to Screen_Prueba for KTP1200 Basic+ PN 17.0.0.0"; PictureOn "Navigates to Screen_Prueba for KTP1200 Basic+ PN 17.0.0.0"
      on Release: ActivateScreen("Screen_Prueba", 0)
   Button "HmiScreenItemData_2" at 36,143 size 159x47; TextOff 'System screens'; PictureOff "Navigates to System screens for KTP1200 Basic+ PN 17.0.0.0"; PictureOn "Navigates to System screens for KTP1200 Basic+ PN 17.0.0.0"
      on Release: ActivateScreen("System screens", 0)

screen "Screen_Prueba" 1280x800, template "Template_1"
   on GenerateScreen: SetTag("Tag_ScreenNumber", 2)
   TextField "HmiScreenItemData" at 128,384 size 1024x27; Text 'Screen_Prueba'
   Button "Back" at 1,49 size 159x47; TextOff 'Back'
      on Release: ActivateScreen("Root screen", 0)